   1285: 'GCU_WARNING_WORD_09_BIT_5', class GCU Warnings, trigger "62_Warning_Data_GCU_WARNING_WORD_09" bit 13
   1286: 'GCU_WARNING_WORD_09_BIT_6', class GCU Warnings, trigger "62_Warning_Data_GCU_WARNING_WORD_09" bit 14
   1287: 'GCU_WARNING_WORD_09_BIT_7', class GCU Warnings, trigger "62_Warning_Data_GCU_WARNING_WORD_09" bit 15
   2384: '', class Tank Control Warnings, trigger "2062_Warning_Data_BTCS_WARNING_WORD_17" bit 0
   2385: '', class Tank Control Warnings, trigger "2062_Warning_Data_BTCS_WARNING_WORD_17" bit 1
   2386: '', class Tank Control Warnings, trigger "2062_Warning_Data_BTCS_WARNING_WORD_17" bit 2
   2387: '', class Tank Control Warnings, trigger "2062_Warning_Data_BTCS_WARNING_WORD_17" bit 3
   2388: '', class Tank Control Warnings, trigger "2062_Warning_Data_BTCS_WARNING_WORD_17" bit 4
   2389: '', class Tank Control Warnings, trigger "2062_Warning_Data_BTCS_WARNING_WORD_17" bit 5
   2390: '', class Tank Control Warnings, trigger "2062_Warning_Data_BTCS_WARNING_WORD_17" bit 6
   2391: '', class Tank Control Warnings, trigger "2062_Warning_Data_BTCS_WARNING_WORD_17" bit 7
   2392: 'DO427 3S OUT OF RANGE', class Tank Control Warnings, trigger "2062_Warning_Data_BTCS_WARNING_WORD_17" bit 8
   2393: 'DO428 4P OUT OF RANGE', class Tank Control Warnings, trigger "2062_Warning_Data_BTCS_WARNING_WORD_17" bit 9
   2394: 'DO427 4S OUT OF RANGE', class Tank Control Warnings, trigger "2062_Warning_Data_BTCS_WARNING_WORD_17" bit 10
   2395: 'DO428 5P OUT OF RANGE', class Tank Control Warnings, trigger "2062_Warning_Data_BTCS_WARNING_WORD_17" bit 11
   2396: 'DO427 5S OUT OF RANGE', class Tank Control Warnings, trigger "2062_Warning_Data_BTCS_WARNING_WORD_17" bit 12
   2397: 'DO428 6P OUT OF RANGE', class Tank Control Warnings, trigger "2062_Warning_Data_BTCS_WARNING_WORD_17" bit 13
   2398: 'DO427 6S OUT OF RANGE', class Tank Control Warnings, trigger "2062_Warning_Data_BTCS_WARNING_WORD_17" bit 14
   2399: 'DO428 APT OUT OF RANGE', class Tank Control Warnings, trigger "2062_Warning_Data_BTCS_WARNING_WORD_17" bit 15

text list "P301 Present": 0..1 'P301 Not Pres'; 1 'P301 Present'

text list "CV312 Present": 0..1 'CV312 Not Pres'; 1 'CV312 Present'

text list "CV431 Present": 0..1 'CV431 Not Pres'; 1 'CV431 Present'

text list "CV432 Present": 0..1 'CV432 Not Pres'; 1 'CV432 Present'

text list "STEP LIST IGG": 1 'Step 001 = Confirm Auto Conditions Ok'; 5 'Step 005 = Wait for Start IGG Command'; 10 'Step 010 = Start E131 (IA Compressor)'; 20 'Step 020 = IA Pressure Within Range (PIT112)'; 30 'Step 030 = CSW Outlet Valves In Position'; 40 'Step 040 = CSW Inlet Valves In Position'; 50 'Step 050 = Start P301 (CSW Pump)'; 60 'Step 060 = CSW Inlet pressure Check'; 70 'Step 070 = Check CV203 Position Closed (N.C.)'; 80 'Step 080 = Start E500 (Fuel Pump)'; 90 'Step 090 = Fuel Pressure Within Range (PIT204)'; 100 'Step 100 = Start E139 (CAB)'; 110 'Step 110 = Start Modulation CV403 (Vent Valve) & Check Setpoint Setting'; 120 'Step 120 = Outlet Pressure Within Range (PIT402)'; 130 'Step 130 = Adjust PIT102 Setpoints'; 140 'Step 140 = Pre BC Start Sequence Delay'; 150 'Step 150 = BC Start Command'; 160 'Step 160 = Wait For Pilot Burner Active Status'; 170 'Step 170 = Adjust Setpoints'; 180 'Step 180 = Wait For Pilot Burner Purge Stage Complete'; 190 'Step 190 = Run Setpoint Ramp For PIT402'; 200 'Step 200 = BC Ramp O2 Command'; 210 'Step 210 = Wait For O2 Level OK'; 220 'Step 220 = Wait For Stop Command'; 300 'Step 300 = Stop Command To BC'; 310 'Step 310 = Wait For Stopping Status From BC'; 320 'Step 320 = Wait For O2 Control Stopped From BC'; 330 'Step 330 = Adjust Setpoints'; 340 'Step 340 = Run Setpoint Ramp Down For PIT402'; 350 'Step 350 = Command Burners Off'; 360 'Step 360 = CV403 To 100% (Fully Open)'; 370 'Step 370 = Adjust Setpoints'; 380 'Step 380 = Stop Combustion Air Blower E139'; 390 'Step 390 = Close CV127 Command To BC'; 400 'Step 400 = Stop Fuel Pump'; 410 'Step 410 = Pre CV203 Close Command Delay'; 420 'Step 420 = Close CV203 Command To BC'; 430 'Step 430 = Stop P301 (CSW Pump)'; 440 'Step 440 = P301 Stopped Delay'; 450 'Step 450 = Cooling Water inlet Valves To Initial Position CV311 = Closed & CV312 = Open'; 460 'Step 460 = CV311 Closed Delay'; 470 'Step 470 = Cooling Water Outlet Valves To Initial Position CV321 = Open & CV322 = Closed'; 480 'Step 480 = CV321 Opened Delay'; 490 'Step 490 = Close CV111 Command To BC'; 500 'Step 500 = Wait For Shutdown Status From BC'

text list "STEP LIST BC": 1 'Step 001 = Confirm Auto Conditions Ok'; 5 'Step 005 = Wait for Start BC Command'; 10 'Step 010 = Open Test Pressure valve CV127'; 20 'Step 020 = Check Pressure PS101'; 30 'Step 030 = CV127 Open Delay #1'; 40 'Step 040 = Check Pressure PS101'; 50 'Step 050 = Close Test Pressure valve CV127'; 60 'Step 060 = Check No Pressure PS101'; 70 'Step 070 = CV127 Closed Delay'; 80 'Step 080 = Check No Pressure PS101'; 90 'Step 090 = Open Test Pressure valve CV127'; 100 'Step 100 = Check Pressure PS101'; 110 'Step 110 = CV127 Open Delay #2'; 120 'Step 120 = Check Pressure PS101'; 130 'Step 130 = Open Pilot Burner Ignition Air Valve CV124'; 140 'Step140 = CV124 Open Delay'; 150 'Step 150 = Check Flow FS123'; 160 'Step 160 = Pilot Flame Ignition Sequence Done OK'; 170 'Step 170 = Wait For IGG Confirmation To Continue'; 180 'Step180 = Open CV114'; 190 'Step 190 = CV114 Open Delay'; 200 'Step 200 = Main Burner Ignition Sequence'; 210 'Step 210 = Check Pressure PIT113'; 220 'Step 220 = Pilot Burner Purge Sequence'; 300 'Step 300 = Confirm Shutting Down'; 310 'Step 310 = CV203 To High O2 Standard Burn Setting'; 320 'Step 320 = CV111 To High O2 Standard Burn Setting'; 330 'Step 330 = Modulation Stopped Confirmation To IGG'; 340 'Step 340 = Wait For Stop Burns Command'; 350 'Step 350 = Close CV206'; 360 'Step 360 = CV206 Close Delay'; 370 'Step 370 = Close CV207'; 380 'Step 380 = CV207 Close Delay'; 390 'Step 390 = Close CV114'; 400 'Step 400 = CV114 Close Delay'; 410 'Step 410 = Close CV215'; 420 'Step 420 = CV215 Close Delay'; 430 'Step 430 = Close CV216'; 440 'Step 440 = CV216 Close Delay'; 450 'Step 450 = Close CV124'; 460 'Step 460 = CV124 Close Delay'; 470 'Step 470 = Check No Flame'; 480 'Step 480 = Burn Stopped Confirmation To IGG'; 490 'Step 490 = Wait For Close CV127 Command'; 500 'Step 500 = Close CV127'; 95 'Step 095 = Confirm CV403 Is Open'; 230 'Step 230 = Wait For Ramp O2 Command'; 240 'Step 240 = Run O2 Ramp'; 250 'Step 250 = Wait For O2 In Specification'; 260 'Step 260 = Write O2 Within Specification Status To IGG'; 270 'Step 270 = Wait For Shutdown Command'; 510 'Step 510 = CV127 Close Delay'; 520 'Step 520 = CV127 Closed Confirmation To IGG'; 525 'Step 525 = Wait For Close CV203 Command'; 530 'Step 530 = Close CV203'; 540 'Step 540 = CV203 Closed Confirmation To IGG'; 550 'Step 550 = Wait For Close CV111 Command'; 560 'Step 560 = Close CV111'; 570 'Step 570 = Shutdown Done Status To IGG'

text list "Mod de functionare motor": 1 'AUTOMATIC PLC'; 0 'LOCAL CABINET'; 2 'MANUAL SCADA'; 3 'MANUAL HMI'; 4 'Necunoscut'

text list "Stari motor": 1 'În pauza de răcire'; 2 'Gata de lucru'; 3 'În functiune'; 4 'În avarie'; 5 'Deconectat'; 6 'Condiţii de start OK'; 7 'Necunoscut'

text list "Mod comanda SP1 Automat": 0 'MANUAL'; 1 'AUTOMATIC'

text list "STATE LIST BTCS": 0 'Initial = Waiting for start'; 1 'Pre-Dwell = Period prior to de-oxygenation'; 2 'De-Ox = De-oxygenation'; 3 'Dwell = Period prior to re-oxygenation'; 4 'Re-Ox = Re-oxygenation'; 5 'Post-Dwell = Settle period'; 6 'Shut Down = System shutting down'

text list "Port Tank": 0 'Deactivated'; 1 'Activated'

text list "STEP LIST BTCS": 0 '00 = Initialising'; 1 '01 = Wait for accept & launch'; 5 '05 = Count to prep gas, 30 Mins from Pre-dwell done'; 10 '10 = Wait for preparing gas confirmation'; 15 '15 = Wait For Pre Dwell Done & Gas Available'; 20 '20 = Close activated tank vent valves'; 25 '25 = Open CV406 Gas to deck valve'; 30 '30 = Open CV407 Block valve 1'; 35 '35 = Open CV411 Block valve 2'; 40 '40 = Close CV409 Blead Valve'; 45 '50 = 15s Time delay'; 50 '50 = Open Activated Tank GTT Valves (Gas To Tank)'; 55 '55 = Wait for O2 @ SP For active tanks for 1 minute'; 60 '60 = Wait For DeOx & DeOx @ SP Times Done'; 70 '70 = Confirm IGG Shutdown'; 75 '75 = Close Activated Tank GTT Valves (Gas To Tank)'; 80 '80 = 30s Time delay'; 85 '85 = Open CV409 Blead Valve'; 90 '90 = Close CV406 Gas to deck valve'; 95 '95 = Close CV407 Block Valve 1'; 100 '100 = Close CV411 Block Valve 2'; 110 '110 = Wait For Dwell Time Done'; 120 '120 = Open All Activated Tank Vent Valves'; 125 '125 = Open CV406 Gas to deck valve'; 130 '130 = Open CV407 Block valve 1'; 135 '135 = Open CV411 Block valve 2'; 140 '140 = Close CV409 Blead Valve'; 145 '150 = 15s Time delay'; 150 '150 = Open Activated Tank GTT Valves (Gas To Tank)'; 155 '155 = Wait for O2 @ SP For active tanks for 1 minute'; 160 '160 = Wait For ReOx & ReOx @ SP Times Done'; 170 '170 = Confirm Gas Deleivery Shutdown'; 175 '175 = Close Activated Tank GTT Valves (Gas To Tank)'; 180 '180 = 30s Time delay'; 185 '185 = Open CV409 Blead Valve'; 190 '190 = Close CV406 Gas to deck valve'; 195 '195 = Close CV407 Block Valve 1'; 200 '200 = Close CV411 Block Valve 2'; 210 '210 = Wait For Dwell Time Done'; 220 '220 = System At Shutdown Goto Initialise'

text list "STEP LIST_GCU": 1 'Step 001 = Confirm Auto Conditions Ok'; 5 'Step 005 = Wait For Tank System State Needing Gas'; 10 'Step 010 = Wait For Prepare Gas Command'; 20 'Step 020 = Run Command To IGG'; 30 'Step 030 = Wait For Running & O2 OK Status From IGG'; 40 'Step 040 = Wait For Supply Gas Command'; 50 'Step 050 = Critical Sensor Check'; 60 'Step 060 = Close CV341'; 70 'Step 070 = CV341 Closed Delay'; 80 'Step 080 = Amend Setpoints'; 90 'Step 090 = Open CV358'; 100 'Step 100 = Start P305 (If Fitted)'; 110 'Step 110 = P305 Started Delay'; 120 'Step 120 = Start P304'; 130 'Step 130 = P304 Started Delay'; 140 'Step 140 = GCU Tank Pre-Fill Delay'; 150 'Step 150 = Fill Sucess Or Fail'; 160 'Step 160 = Stop P304'; 170 'Step 170 = P304 Stopped Delay'; 180 'Step 180 = Stop P305 (If Fitted)'; 190 'Step 190 = P305 Stopped Delay'; 200 'Step 200 = Close CV358'; 210 'Step 210 = CV358 Closed Delay'; 220 'Step 220 = Amend Setpoints'; 230 'Step 230 = Start P303'; 240 'Step 240 = P303 Started Delay'; 250 'Step 250 = Confirm No Alarms'; 260 'Step 260 = Start E400'; 270 'Step 270 = E400 Into Loaded Before Step Time Out (E400 Started Delay)'; 280 'Step 280 = E400 On Load Running Delay'; 290 'Step 290 = CV405 Modulation Start & PIT416 Target Ramp Run'; 300 'Step 300 = Amend Setpoints (Not Currently Required = Re-Check)'; 310 'Step 310 = Wiat For BWTS Status (2=DeOx) or (3=Dwell/ReOx)'; 320 'Step 320 = Open CV401'; 330 'Step 330 = CV401 Opened Delay'; 340 'Step 340 = Pre-Open CV441 Sequence Delay'; 350 'Step 350 = Close CV441'; 360 'Step 360 = CV441 Closed Delay (Done = Jump To Step 410)'; 370 'Step 370 = Close CV401'; 380 'Step 380 = CV401 Closed Delay'; 390 'Step 390 = Open CV441'; 400 'Step 400 = CV441 Opened Delay'; 410 'Step 410 = DeOx/ReOx Valave Configuration Done Sequence Delay'; 420 'Step 420 = Wait For Shutdown Instruction +++RUNNING+++'; 430 'Step 430 = Spare Step (Not Used)'; 440 'Step 440 = Spare Step (Not Used)'; 450 'Step 450 = Open CV405 (Start Of Shutdwon Sequence)'; 460 'Step 460 = CV405 Opened Delay'; 470 'Step 470 = Check CV406 Closed (BWT Control)'; 480 'Step 480 = CV406 Closed Delay'; 490 'Step 490 = Open CV441'; 500 'Step 500 = CV441 Opened Delay'; 510 'Step 510 = Close CV401'; 520 'Step 520 = CV401 Closed Delay'; 530 'Step 530 = Stop E400'; 540 'Step 540 = Stop P303'; 550 'Step 550 = P303 Stopped Delay'; 560 'Step 560 = Wait For PIT416 <0.01bar'; 570 'Step 570 = Open CV341'; 580 'Step 580 = CV341 Opened Delay'; 590 'Step 590 = Tank Drain Time Delay'; 600 'Step 600 = Tank Flush Sequence'; 610 'Step 610 = Post Flush Delay'

text list "P305 Present": 0..1 'P305 Not Pres'; 1 'P305 Present'

text list "GCU_LCL": 0 'TAKE CONTROL'; 1 'RELEASE CONTROL'

text list "ENBL_DSBL": 0 'Disabled'; 1 'Enabled'

text list "GTT_OPS": 0 'Open Active GTT Valves'; 1 'Close Active GTT Valves'

text list "BTCS/BWTC": 0 'Activate'; 1 'Deactivate'

text list "PGC Commissioning": 0 'MEA Tank Changeover'; 1 'Please Wait'

text list "IG Transfer": 0 'Cargo Blanketing Mode'; 1 'Balast Water Treatment Mode'

text list "m³/hr to Nm³/hr": 0 'm³/hr to Nm³/hr Conversion'; 1 'm³/hr Raw Value'

graphic list "IA Compressor": 3 'IA Compressor 01'; 0 'IA Compressor 01'; 1 'IA Compressor 02_1'; 2 'IA Compressor 0_1'

graphic list "New IA Compressor": 0 'Graphic_249'; 1 'Graphic_250'; 2 'Graphic_249'; 3 'Graphic_250'

graphic list "Pump Ani": 1 'Pumpd'; 0 'Pump0'; 1 'Pump1'; 2 'Pump2'; 5 'Pumpd'; 3 'Pump0'; 4 'Pump1'

graphic list "IA Compressor_1": 3 'IA Compressor 01'; 0 'IA Compressor 0_1'; 1 'IA Compressor 02_1'; 2 'IA Compressor 0_1'; 0 'IA Compressor 01'

graphic list "IA Compressor_2": 3 'IA Compressor 01'; 0 'IA Compressor 0_1'; 1 'IA Compressor 02_1'; 2 'IA Compressor 0_1'; 0 'IA Compressor 01'

graphic list "IGGS": 0 'Graphic_3'; 1 'Graphic_140'

graphic list "GCU": 0 'Graphic_150'; 1 'Graphic_150'

graphic list "Process time Banner": 2..5 'Graphic_193'; 1 'Pre Dwell'; 2 'Graphic_193'

graphic list "Tank Process Stage_II": 0 'INITIAL STATE'; 1 'Pre Dwell'; 2 'De-Oxygenation'; 3 'Graphic_189'; 4 'Graphic_190'; 5 'Graphic_191'; 6 'Graphic_192'; 7 'Graphic_186'

graphic list "Water Level Override": 0 'Graphic_217'; 1 'Graphic_218'; 2 'Graphic_217'

graphic list "LED": 0 'PilotLight_Round_G_Off_256c'; 1 'PilotLight_Round_G_On_256c'

Template "Template" 1280x800
   Button "HmiScreenItemData_12" at 953,4 size 80x35; TextOn 'WARNING'; TextOff 'Warning'
      on Release: ActivateScreen("04 Alarm Log", 0)
      Visibility <- "62_Warning_Data_WRNG_PRSNT"
   Button "HmiScreenItemData_14" at 1040,4 size 80x35; TextOn 'ALARM'; TextOff 'Alarm'
      on Release: ActivateScreen("04 Alarm Log", 0)
      Visibility <- "60_Alarm_Data_ALRM_PRSNT"
   Button "HmiScreenItemData_20" at 866,4 size 80x35; TextOn 'Back'; TextOff 'Lockout'
      on Click: SetBit("80_From_HMI_Reset_Alarms")
      on Press: function_b14e0dd5("80_From_HMI_RST_LOCKOUT", 0)
      Appearance <- "82_To_HMI_E-STOP LATCHED"
   Button "HmiScreenItemData_24" at 770,3 size 64x35; TextOn 'MUTE'; TextOff 'Mute'
      on Press: function_b14e0dd5("80_From_HMI_SLNCE_BZR", 0)
      Appearance <- "80_From_HMI_SLNCE_BZR"
   GraphicView "Graphic view_24" at 836,3 size 29x41; Picture "Graphic_138"
      Visibility <- "Buzzer"
   Group "Group_11" at 300,4 size 240x30
   Button "HmiScreenItemData_26" at 547,4 size 216x31; TextOn 'Back'; TextOff 'Text'
   IOField "I/O field_9" at 636,8 size 40x23; FormatPattern 99; Unit h
      ProcessValue <- "103_Main_Burner_DB_Hours burn_CV"
   IOField "I/O field_16" at 677,8 size 40x23; FormatPattern 99; Unit m
      ProcessValue <- "103_Main_Burner_DB_Minutes burn_CV"
   IOField "I/O field_19" at 718,8 size 40x23; FormatPattern 99; Unit s
      ProcessValue <- "103_Main_Burner_DB_Seconds burn_CV"
   GraphicView "Graphic view_80" at 544,-4 size 59x52; Picture "Graphic_130"
      Visibility <- "103_Main_Burner_DB_DN_OK"
   IOField "I/O field_35" at 595,8 size 40x23; FormatPattern 99; Unit d
      ProcessValue <- "103_Main_Burner_DB_Days burn_CV"
   Circle "Circle_46" at 265,6 size 26x26
      Appearance <- "IGG PLC HEART BEAT"
      Visibility <- "TRUE"
   Circle "Circle_1" at 235,6 size 26x26
      Visibility <- "TRUE"
      Appearance <- "Setpoint Override_DB_Set Pressure"
   Button "Button_8" at 300,4 size 240x30; TextOn 'IGGS Shutting Down'; TextOff 'IGGS Shutting down'
      Visibility <- "100_IGG_AUTO_SEQ_DB_CRNT_STEP"
   Button "Button_2" at 300,4 size 240x30; TextOn 'IGGS Starting Up'; TextOff 'IGGS Starting Up'
      Visibility <- "100_IGG_AUTO_SEQ_DB_CRNT_STEP"

screen "01 Home" 1280x800, template "Template"
   GraphicView "Graphic view_2" at 118,52 size 317x684; Picture "Graphic_137"
   TextField "HmiScreenItemData_4" at 204,164 size 865x50; Text 'Welcome to Coldharbour Marine'
   TextField "HmiScreenItemData_3" at 194,220 size 896x88; Text 'Ballast Water Treatment System'
   Button "HmiScreenItemData" at 116,50 size 1048x686; TextOn 'Main Index'; TextOff 'Text'
      on Release: function_a2a04561(); ActivateScreen("02 Main Index", 0)
   GraphicView "Graphic view_1" at 444,350 size 449x266; Picture "Graphic_185"
   Button "HmiScreenItemData_16" at 98,47 size 1089x692; TextOn 'Back'; TextOff 'Text'
      on Release: function_a2a04561(); ActivateScreen("Balast Water Treatment Plant", 0)
   Button "Button_1" at 1222,758 size 56x40; TextOff 'Text'; PictureOff "Graphic_286"; Authorization "User administration"
      on Release: StopRuntime(0)

screen "03 User Admin" 1280x800, template "Template"
   Button "HmiScreenItemData_1" at 1,1 size 159x51; TextOn 'Back'; TextOff 'Main Index'
      on Release: ActivateScreen("02 Main Index", 0)
   UserView "User view_1" at 0,69 size 1279x730
   Button "HmiScreenItemData_4" at 1153,16 size 126x33; TextOn 'I&A Compressor Ok'; TextOff 'Previous Screen'
      on Release: function_efd93a16()

screen "05 Alarm Buffer" 1280x800, template "Template"
   AlarmView "Alarm view_1" at 8,61 size 1258x729
   Button "HmiScreenItemData_2" at 143,2 size 139x43; TextOn 'Back'; TextOff 'Alarm'
      on Release: ActivateScreen("04 Alarm Log", 0)
   Button "HmiScreenItemData_5" at 1,2 size 139x43; TextOn 'Back'; TextOff 'Main Index'
      on Release: ActivateScreen("02 Main Index", 0)
   Button "HmiScreenItemData_4" at 1138,1 size 139x43; TextOn 'I&A Compressor Ok'; TextOff 'Back'
      on Release: function_efd93a16()

screen "07 BWTS MAIN" 1280x800, template "Template"
   Rectangle "Rectangle_2" at 150,205 size 480x40
      Appearance <- "2102_TIME_CALCS_DB_DE_OX_TMR_DN"
   TextField "Text field_7" at 155,210 size 200x30; Text 'De-Oxygenate Time :'
   IOField "I/O field_3" at 360,210 size 60x30; FormatPattern 999
      ProcessValue <- "2110_BTCS_CNTRL_DB_DE_OX_HRS"
   TextField "Text field_8" at 420,210 size 60x30; Text 'Hours'
   IOField "I/O field_4" at 485,210 size 60x30; FormatPattern 99
      ProcessValue <- "2110_BTCS_CNTRL_DB_DE_OX_MINS"
   TextField "Text field_9" at 545,210 size 80x30; Text 'Minutes'
   Rectangle "Rectangle_3" at 150,250 size 480x40
      Appearance <- "2102_TIME_CALCS_DB_DWELL_TMR_DN"
   TextField "Text field_10" at 155,255 size 200x30; Text 'Dwell Time :'
   IOField "I/O field_5" at 360,255 size 60x30; FormatPattern 999
      ProcessValue <- "2110_BTCS_CNTRL_DB_DWELL_HRS"
   TextField "Text field_11" at 420,255 size 60x30; Text 'Hours'
   IOField "I/O field_6" at 485,255 size 60x30; FormatPattern 99
      ProcessValue <- "2110_BTCS_CNTRL_DB_DWELL_MINS"
   TextField "Text field_12" at 545,255 size 80x30; Text 'Minutes'
   Rectangle "Rectangle_4" at 150,295 size 480x40
      Appearance <- "2102_TIME_CALCS_DB_RE_OX_TMR_DN"
   TextField "Text field_13" at 155,300 size 200x30; Text 'Re-Oxygenate Time :'
   IOField "I/O field_7" at 360,300 size 60x30; FormatPattern 999
      ProcessValue <- "2110_BTCS_CNTRL_DB_RE_OX_HRS"
   TextField "Text field_14" at 420,300 size 60x30; Text 'Hours'
   IOField "I/O field_8" at 485,300 size 60x30; FormatPattern 99
      ProcessValue <- "2110_BTCS_CNTRL_DB_RE_OX_MINS"
   TextField "Text field_15" at 545,300 size 80x30; Text 'Minutes'
   Rectangle "Rectangle_5" at 150,340 size 480x40
      Appearance <- "2102_TIME_CALCS_DB_POST_DWELL_TMR_DN"
   TextField "Text field_16" at 155,345 size 200x30; Text 'Post-Dwell Time :'
   IOField "I/O field_9" at 360,345 size 60x30; FormatPattern 999
      ProcessValue <- "2110_BTCS_CNTRL_DB_POST_DWELL_HRS"
   TextField "Text field_17" at 420,345 size 60x30; Text 'Hours'
   IOField "I/O field_10" at 485,345 size 60x30; FormatPattern 99
      ProcessValue <- "2110_BTCS_CNTRL_DB_POST_DWELL_MINS"
   TextField "Text field_18" at 545,345 size 80x30; Text 'Minutes'
   Rectangle "Rectangle_6" at 640,205 size 480x40
      Appearance <- "2102_TIME_CALCS_DB_DE_OX_SP_TMR_DN"
   TextField "Text field_19" at 645,210 size 200x30; Text 'At De-Ox Setpoint :'
   IOField "I/O field_11" at 850,210 size 60x30; FormatPattern 999
      ProcessValue <- "2110_BTCS_CNTRL_DB_DE_OX_SP_HRS"
   TextField "Text field_20" at 910,210 size 60x30; Text 'Hours'
   IOField "I/O field_12" at 975,210 size 60x30; FormatPattern 99
      ProcessValue <- "2110_BTCS_CNTRL_DB_DE_OX_SP_MINS"
   TextField "Text field_21" at 1035,210 size 80x30; Text 'Minutes'
   Rectangle "Rectangle_7" at 640,295 size 480x40
      Appearance <- "2102_TIME_CALCS_DB_RE_OX_SP_TMR_DN"
   TextField "Text field_22" at 645,300 size 200x30; Text 'At Re-Ox Setpoint :'
   IOField "I/O field_13" at 850,300 size 60x30; FormatPattern 999
      ProcessValue <- "2110_BTCS_CNTRL_DB_RE_OX_SP_HRS"
   TextField "Text field_23" at 910,300 size 60x30; Text 'Hours'
   IOField "I/O field_14" at 975,300 size 60x30; FormatPattern 99
      ProcessValue <- "2110_BTCS_CNTRL_DB_RE_OX_SP_MINS"
   TextField "Text field_24" at 1035,300 size 80x30; Text 'Minutes'
   TextField "Text field_25" at 155,435 size 200x30; Text 'Total Sequence Time:'
   IOField "I/O field_15" at 360,435 size 60x30; FormatPattern 999
      ProcessValue <- "2110_BTCS_CNTRL_DB_TOT_SEQ_HRS"
   TextField "Text field_26" at 420,435 size 60x30; Text 'Hours'
   IOField "I/O field_16" at 485,435 size 60x30; FormatPattern 99
      ProcessValue <- "2110_BTCS_CNTRL_DB_TOT_SEQ_MINS"
   TextField "Text field_27" at 545,435 size 80x30; Text 'Minutes'
   TextField "Text field_28" at 155,625 size 200x30; Text 'Remaining Time:'
   IOField "I/O field_17" at 360,625 size 60x30; FormatPattern 999
      ProcessValue <- "2110_BTCS_CNTRL_DB_RMNG_SEQ_HRS"
   TextField "Text field_29" at 420,625 size 60x30; Text 'Hours'
   IOField "I/O field_18" at 485,625 size 60x30; FormatPattern 99
      ProcessValue <- "2110_BTCS_CNTRL_DB_RMNG_SEQ_MINS"
   TextField "Text field_30" at 545,625 size 80x30; Text 'Minutes'
   Button "HmiScreenItemData_1" at 10,10 size 160x50; TextOn 'Back'; TextOff 'Main Index'
      on Release: ActivateScreen("02 Main Index", 0)
   TextField "Text field_1" at 320,10 size 640x35; Text 'BASIC BARGE TWO TANK CONTROL SYSTEM'
   Button "HmiScreenItemData_2" at 1110,10 size 160x50; TextOn 'Back'; TextOff 'Enable'
      on Press: ResetBit("80_From_HMI_RUN_BWTS"); SetBit("80_From_HMI_RUN_BTCS")
      Visibility <- "80_From_HMI_RUN_BWTS"
   Button "HmiScreenItemData_3" at 918,75 size 160x50; TextOn 'Back'; TextOff 'Disable'
      on Press: ResetBit("80_From_HMI_RUN_BTCS"); SetBit("80_From_HMI_RUN_BWTS")
      Visibility <- "80_From_HMI_RUN_BTCS"
   TextField "Text field_2" at 480,40 size 320x35; Text 'BTCS ENABLED'
      Visibility <- "80_From_HMI_RUN_BTCS"
   TextField "Text field_3" at 480,40 size 320x35; Text 'BTCS DISABLED'
      Visibility <- "80_From_HMI_RUN_BTCS"
   Button "Button_2" at 10,70 size 160x50; TextOn 'User Account'; TextOff 'Alarm Log'; Authorization "User administration"
      on Release: ActivateScreen("04 Alarm Log", 0)
   Group "Group_1" at 150,205 size 480x40
   Group "Group_2" at 150,250 size 480x40
   Group "Group_3" at 150,295 size 480x40
   Group "Group_4" at 150,340 size 480x40
   Group "Group_5" at 640,205 size 480x40
   Group "Group_6" at 640,295 size 480x40
   Group "Group_7" at 150,430 size 480x40
   Group "Group_8" at 150,620 size 480x40
   TextField "Text field_31" at 1005,150 size 120x30; Text 'SETUP'
   TextField "Text field_32" at 1005,420 size 120x30; Text 'CONTROL'
   Button "Button_1" at 150,520 size 230x50; TextOff 'ACCEPT & LAUNCH'
      on Release: ResetBit("2110_BTCS_CNTRL_DB_START_SEQ")
      on Press: SetBit("2110_BTCS_CNTRL_DB_START_SEQ")
      Appearance <- "2110_BTCS_CNTRL_DB_BTCS_STATE"
      Visibility <- "2102_TIME_CALCS_DB_TIMES_VALID"
   SymbolicIOField "Symbolic I/O field_1" at 640,480 size 480x30; TextOn '1'; TextOff '0'; TextList "STATE LIST BTCS"
      ProcessValue <- "2110_BTCS_CNTRL_DB_BTCS_STATE"
   TextField "Text field_33" at 150,480 size 480x35; Text 'TIMES NOT VALID'
      Visibility <- "2102_TIME_CALCS_DB_TIMES_VALID"
   TextField "Text field_34" at 150,480 size 480x35; Text 'TIMES VALID'
      Visibility <- "2102_TIME_CALCS_DB_TIMES_VALID"
   SymbolicIOField "Symbolic I/O field_2" at 640,580 size 480x30; TextOn '1'; TextOff '0'; TextList "STEP LIST BTCS"
      ProcessValue <- "2110_BTCS_CNTRL_DB_BTCS_STEP"
   Button "HmiScreenItemData_4" at 1110,70 size 160x50; TextOn 'Back'; TextOff 'Master Reset'
      on Press: ResetBit("2110_BTCS_CNTRL_DB_RESET_ALL"); SetBit("2110_BTCS_CNTRL_DB_RESET_ALL")
      Visibility <- "80_From_HMI_RUN_BTCS"
   SymbolicIOField "Symbolic I/O field_3" at 360,700 size 140x30; TextOn '1'; TextOff '0'; TextList "Port Tank"
      ProcessValue <- "2110_BTCS_CNTRL_DB_PORT_TANK_STS"
   Button "Button_4" at 150,700 size 180x30; TextOff 'Port Tank'
      on Press: InvertBit("2110_BTCS_CNTRL_DB_PORT_TANK_STS")
      Appearance <- "2110_BTCS_CNTRL_DB_PORT_TANK_STS"
   TextField "Text field_35" at 1025,690 size 100x30; Text 'TANKS'
   SymbolicIOField "Symbolic I/O field_4" at 360,740 size 140x30; TextOn '1'; TextOff '0'; TextList "Port Tank"
      ProcessValue <- "2110_BTCS_CNTRL_DB_STBD_TANK_STS"
   Button "Button_5" at 150,740 size 180x30; TextOff 'Starboard Tank'
      on Press: InvertBit("2110_BTCS_CNTRL_DB_STBD_TANK_STS")
      Appearance <- "2110_BTCS_CNTRL_DB_STBD_TANK_STS"
   TextField "Text field_37" at 515,700 size 60x30; Text 'O2 :'
   IOField "I/O field_20" at 575,700 size 60x30; FormatPattern 99.99
      ProcessValue <- "20_TANKS_IP_DATA_RIO_02_FIRST_TANK_BWT_DO"
   TextField "Text field_36" at 640,700 size 60x30; Text 'ph :'
   IOField "I/O field_19" at 700,700 size 60x30; FormatPattern 99.99
      ProcessValue <- "20_TANKS_IP_DATA_RIO_02_FIRST_TANK_BWT_PH"
   TextField "Text field_38" at 775,700 size 65x30; Text 'Temp :'
   IOField "I/O field_21" at 840,700 size 60x30; FormatPattern 99.99
      ProcessValue <- "20_TANKS_IP_DATA_RIO_02_FIRST_TANK_BWT_TEMP"
   TextField "Text field_39" at 910,700 size 65x30; Text 'Level :'
   IOField "I/O field_22" at 975,700 size 60x30; FormatPattern 99.9
      ProcessValue <- "20_TANKS_IP_DATA_RIO_02_FIRST_TANK_BWT_LEVEL"
   TextField "Text field_40" at 515,740 size 60x30; Text 'O2 :'
   IOField "I/O field_23" at 575,740 size 60x30; FormatPattern 99.99
      ProcessValue <- "20_TANKS_IP_DATA_RIO_02_SECOND_TANK_BWT_DO"
   TextField "Text field_41" at 640,740 size 60x30; Text 'ph :'
   IOField "I/O field_24" at 700,740 size 60x30; FormatPattern 99.99
      ProcessValue <- "20_TANKS_IP_DATA_RIO_02_SECOND_TANK_BWT_PH"
   TextField "Text field_42" at 775,740 size 65x30; Text 'Temp :'
   IOField "I/O field_25" at 840,740 size 60x30; FormatPattern 99.99
      ProcessValue <- "20_TANKS_IP_DATA_RIO_02_SECOND_TANK_BWT_TEMP"
   TextField "Text field_43" at 910,740 size 65x30; Text 'Level :'
   IOField "I/O field_26" at 975,740 size 60x30; FormatPattern 99.9
      ProcessValue <- "20_TANKS_IP_DATA_RIO_02_SECOND_TANK_BWT_LEVEL"
   Group "Group" at 150,160 size 480x40
   Group "Group_9" at 150,160 size 480x40
   Group "Group_10" at 150,340 size 480x40
   Group "Group_12" at 150,295 size 480x40
   Group "Group_13" at 640,205 size 480x40
   Group "Group_14" at 150,250 size 480x40
   Group "Group_15" at 150,205 size 480x40
   Group "Group_16" at 640,295 size 480x40
   Rectangle "Rectangle_15" at 150,480 size 480x130
      Visibility <- "2100_AUTO_SEQ_DB_SEQ_RNG"
   Button "Button_3" at 400,520 size 230x50; TextOff 'ABORT - STOP'
      on Release: ResetBit("2110_BTCS_CNTRL_DB_STOP_SEQ")
      on Press: SetBit("2110_BTCS_CNTRL_DB_STOP_SEQ")
      Appearance <- "2110_BTCS_CNTRL_DB_BTCS_STATE"
   TextField "Text field_48" at 23,309 size 1188x123; Text 'Re - Work Required Througout This page'
   Rectangle "Rectangle_1" at 150,160 size 480x40
      Appearance <- "2102_TIME_CALCS_DB_PRE_DWELL_TMR_DN"
   TextField "Text field_4" at 155,165 size 200x30; Text 'Pre-Dwell Time :'
   IOField "I/O field_1" at 360,165 size 60x30; FormatPattern 999
      ProcessValue <- "2110_BTCS_CNTRL_DB_PRE_DWELL_HRS"
   TextField "Text field_5" at 420,165 size 60x30; Text 'Hours'
   IOField "I/O field_2" at 485,165 size 60x30; FormatPattern 99
      ProcessValue <- "2110_BTCS_CNTRL_DB_PRE_DWELL_MINS"
   TextField "Text field_6" at 545,165 size 80x30; Text 'Minutes'
   Rectangle "Rectangle_13" at 150,160 size 480x40
      Visibility <- "2100_AUTO_SEQ_DB_SEQ_RNG"
      Appearance <- "2102_TIME_CALCS_DB_PRE_DWELL_TMR_DN"
   TextField "Text field_44" at 155,165 size 310x30; Text 'Pre-Dwell Time Remaining :'
      Visibility <- "2100_AUTO_SEQ_DB_SEQ_RNG"
   IOField "I/O field_28" at 465,165 size 80x30; FormatPattern 999999
      ProcessValue <- "2102_TIME_CALCS_DB_PRE_DWELL_MINS_RMNG"
      Visibility <- "2100_AUTO_SEQ_DB_SEQ_RNG"
   TextField "Text field_46" at 545,165 size 80x30; Text 'Minutes'
      Visibility <- "2100_AUTO_SEQ_DB_SEQ_RNG"
   Rectangle "Rectangle_14" at 150,340 size 480x40
      Visibility <- "2100_AUTO_SEQ_DB_SEQ_RNG"
      Appearance <- "2102_TIME_CALCS_DB_POST_DWELL_TMR_DN"
   TextField "Text field_45" at 155,345 size 310x30; Text 'Post-Dwell Time Remaining :'
      Visibility <- "2100_AUTO_SEQ_DB_SEQ_RNG"
   IOField "I/O field_27" at 465,345 size 80x30; FormatPattern 999999
      Visibility <- "2100_AUTO_SEQ_DB_SEQ_RNG"
      ProcessValue <- "2102_TIME_CALCS_DB_POST_DWELL_MINS_RMNG"
   TextField "Text field_47" at 545,345 size 80x30; Text 'Minutes'
      Visibility <- "2100_AUTO_SEQ_DB_SEQ_RNG"
   Rectangle "Rectangle_16" at 150,295 size 480x40
      Visibility <- "2100_AUTO_SEQ_DB_SEQ_RNG"
      Appearance <- "2102_TIME_CALCS_DB_RE_OX_TMR_DN"
   TextField "Text field_50" at 155,300 size 310x30; Text 'Re-Oxygenate Time Remaining :'
      Visibility <- "2100_AUTO_SEQ_DB_SEQ_RNG"
   IOField "I/O field_30" at 465,300 size 80x30; FormatPattern 999999
      Visibility <- "2100_AUTO_SEQ_DB_SEQ_RNG"
      ProcessValue <- "2102_TIME_CALCS_DB_RE_OX_MINS_RMNG"
   TextField "Text field_51" at 545,300 size 80x30; Text 'Minutes'
      Visibility <- "2100_AUTO_SEQ_DB_SEQ_RNG"
   Rectangle "Rectangle_17" at 640,205 size 480x40
      Visibility <- "2100_AUTO_SEQ_DB_SEQ_RNG"
      Appearance <- "2102_TIME_CALCS_DB_DE_OX_SP_TMR_DN"
   TextField "Text field_52" at 645,210 size 310x30; Text 'At De-Ox Time Remaining :'
      Visibility <- "2100_AUTO_SEQ_DB_SEQ_RNG"
   IOField "I/O field_31" at 955,210 size 80x30; FormatPattern 999999
      Visibility <- "2100_AUTO_SEQ_DB_SEQ_RNG"
      ProcessValue <- "2102_TIME_CALCS_DB_DE_OX_SP_MINS_RMNG"
   TextField "Text field_53" at 1035,210 size 80x30; Text 'Minutes'
      Visibility <- "2100_AUTO_SEQ_DB_SEQ_RNG"
   Rectangle "Rectangle_18" at 150,250 size 480x40
      Visibility <- "2100_AUTO_SEQ_DB_SEQ_RNG"
      Appearance <- "2102_TIME_CALCS_DB_DWELL_TMR_DN"
   TextField "Text field_54" at 155,255 size 310x30; Text 'Dwell Time Remaining :'
      Visibility <- "2100_AUTO_SEQ_DB_SEQ_RNG"
   IOField "I/O field_32" at 465,255 size 80x30; FormatPattern 999999
      Visibility <- "2100_AUTO_SEQ_DB_SEQ_RNG"
      ProcessValue <- "2102_TIME_CALCS_DB_DWELL_MINS_RMNG"
   TextField "Text field_55" at 545,255 size 80x30; Text 'Minutes'
      Visibility <- "2100_AUTO_SEQ_DB_SEQ_RNG"
   Rectangle "Rectangle_19" at 150,205 size 480x40
      Visibility <- "2100_AUTO_SEQ_DB_SEQ_RNG"
      Appearance <- "2102_TIME_CALCS_DB_DE_OX_TMR_DN"
   TextField "Text field_56" at 155,210 size 310x30; Text 'De-Oxygenate Time Remaining :'
      Visibility <- "2100_AUTO_SEQ_DB_SEQ_RNG"
   IOField "I/O field_33" at 465,210 size 80x30; FormatPattern 999999
      Visibility <- "2100_AUTO_SEQ_DB_SEQ_RNG"
      ProcessValue <- "2102_TIME_CALCS_DB_DE_OX_MINS_RMNG"
   TextField "Text field_57" at 545,210 size 80x30; Text 'Minutes'
      Visibility <- "2100_AUTO_SEQ_DB_SEQ_RNG"
   Rectangle "Rectangle_20" at 640,295 size 480x40
      Visibility <- "2100_AUTO_SEQ_DB_SEQ_RNG"
      Appearance <- "2102_TIME_CALCS_DB_RE_OX_SP_TMR_DN"
   TextField "Text field_58" at 645,300 size 310x30; Text 'At Re-Ox Time Remaining :'
      Visibility <- "2100_AUTO_SEQ_DB_SEQ_RNG"
   IOField "I/O field_34" at 955,300 size 80x30; FormatPattern 999999
      Visibility <- "2100_AUTO_SEQ_DB_SEQ_RNG"
      ProcessValue <- "2102_TIME_CALCS_DB_RE_OX_SP_MINS_RMNG"
   TextField "Text field_59" at 1035,300 size 80x30; Text 'Minutes'
      Visibility <- "2100_AUTO_SEQ_DB_SEQ_RNG"

